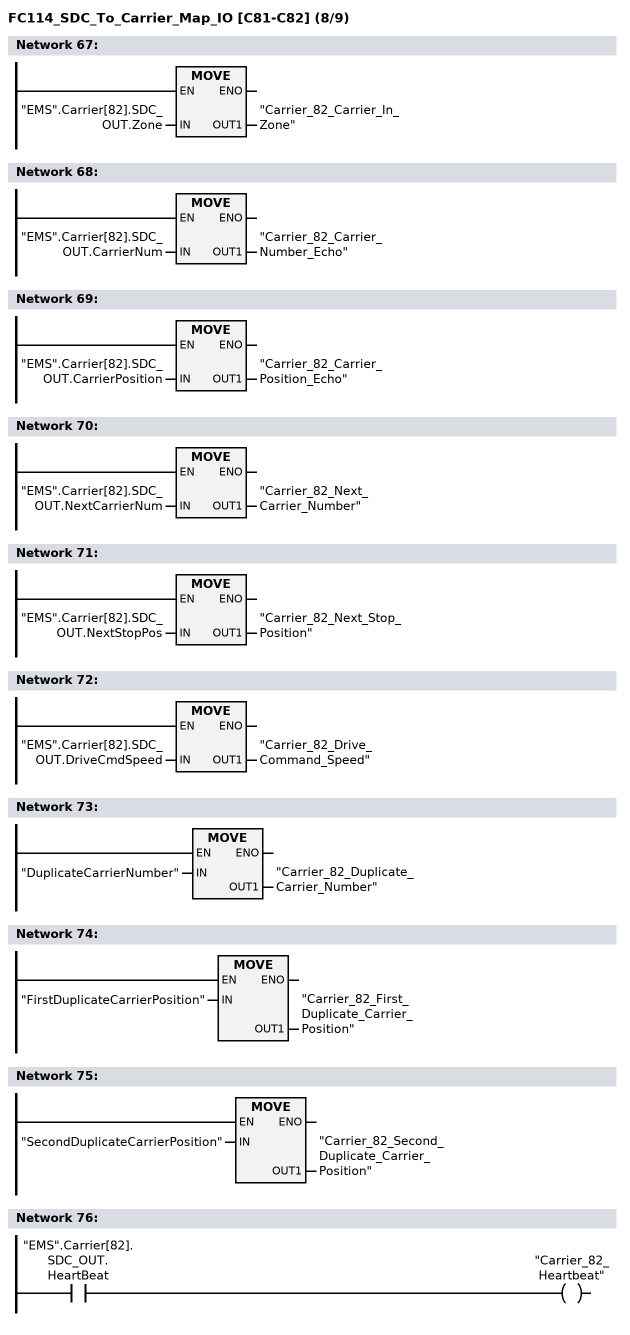
   RUNG wire#powerrail
      Move(in := "EMS".Carrier[82].SDC_OUT.Zone, out1 => "Carrier_82_Carrier_In_Zone")
   END_RUNG
   // the same network as SCL:
   "Carrier_82_Carrier_In_Zone" := "EMS".Carrier[82].SDC_OUT.Zone;
END_REGION

REGION Network 68
   RUNG wire#powerrail
      Move(in := "EMS".Carrier[82].SDC_OUT.CarrierNum, out1 => "Carrier_82_Carrier_Number_Echo")
   END_RUNG
   // the same network as SCL:
   "Carrier_82_Carrier_Number_Echo" := "EMS".Carrier[82].SDC_OUT.CarrierNum;
END_REGION

REGION Network 69
   RUNG wire#powerrail
      Move(in := "EMS".Carrier[82].SDC_OUT.CarrierPosition, out1 => "Carrier_82_Carrier_Position_Echo")
   END_RUNG
   // the same network as SCL:
   "Carrier_82_Carrier_Position_Echo" := "EMS".Carrier[82].SDC_OUT.CarrierPosition;
END_REGION

REGION Network 70
   RUNG wire#powerrail
      Move(in := "EMS".Carrier[82].SDC_OUT.NextCarrierNum, out1 => "Carrier_82_Next_Carrier_Number")
   END_RUNG
   // the same network as SCL:
   "Carrier_82_Next_Carrier_Number" := "EMS".Carrier[82].SDC_OUT.NextCarrierNum;
END_REGION

REGION Network 71
   RUNG wire#powerrail
      Move(in := "EMS".Carrier[82].SDC_OUT.NextStopPos, out1 => "Carrier_82_Next_Stop_Position")
   END_RUNG
   // the same network as SCL:
   "Carrier_82_Next_Stop_Position" := "EMS".Carrier[82].SDC_OUT.NextStopPos;
END_REGION

REGION Network 72
   RUNG wire#powerrail
      Move(in := "EMS".Carrier[82].SDC_OUT.DriveCmdSpeed, out1 => "Carrier_82_Drive_Command_Speed")
   END_RUNG
   // the same network as SCL:
   "Carrier_82_Drive_Command_Speed" := "EMS".Carrier[82].SDC_OUT.DriveCmdSpeed;
END_REGION

REGION Network 73
   RUNG wire#powerrail
      Move(in := "DuplicateCarrierNumber", out1 => "Carrier_82_Duplicate_Carrier_Number")
   END_RUNG
   // the same network as SCL:
   "Carrier_82_Duplicate_Carrier_Number" := "DuplicateCarrierNumber";
END_REGION

REGION Network 74
   RUNG wire#powerrail
      Move(in := "FirstDuplicateCarrierPosition", out1 => "Carrier_82_First_Duplicate_Carrier_Position")
   END_RUNG
   // the same network as SCL:
   "Carrier_82_First_Duplicate_Carrier_Position" := "FirstDuplicateCarrierPosition";
END_REGION

REGION Network 75
   RUNG wire#powerrail
      Move(in := "SecondDuplicateCarrierPosition", out1 => "Carrier_82_Second_Duplicate_Carrier_Position")
   END_RUNG
   // the same network as SCL:
   "Carrier_82_Second_Duplicate_Carrier_Position" := "SecondDuplicateCarrierPosition";
END_REGION

REGION Network 76
   RUNG wire#powerrail
      Contact( "EMS".Carrier[82].SDC_OUT.HeartBeat )
      Coil( "Carrier_82_Heartbeat" )
   END_RUNG
   // the same network as SCL:
   "Carrier_82_Heartbeat" := "EMS".Carrier[82].SDC_OUT.HeartBeat;
END_REGION

REGION Network 77
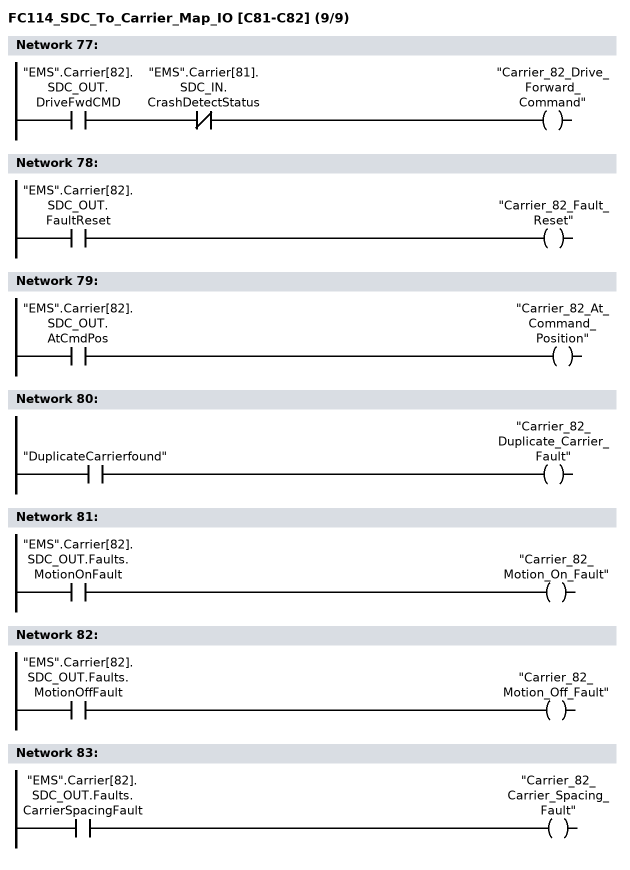
   RUNG wire#powerrail
      Contact( "EMS".Carrier[82].SDC_OUT.DriveFwdCMD )
      I_Contact( "EMS".Carrier[81].SDC_IN.CrashDetectStatus )
      Coil( "Carrier_82_Drive_Forward_Command" )
   END_RUNG
   // the same network as SCL:
   "Carrier_82_Drive_Forward_Command" := "EMS".Carrier[82].SDC_OUT.DriveFwdCMD AND NOT "EMS".Carrier[81].SDC_IN.CrashDetectStatus;
END_REGION

REGION Network 78
   RUNG wire#powerrail
      Contact( "EMS".Carrier[82].SDC_OUT.FaultReset )
      Coil( "Carrier_82_Fault_Reset" )
   END_RUNG
   // the same network as SCL:
   "Carrier_82_Fault_Reset" := "EMS".Carrier[82].SDC_OUT.FaultReset;
END_REGION

REGION Network 79
   RUNG wire#powerrail
      Contact( "EMS".Carrier[82].SDC_OUT.AtCmdPos )
      Coil( "Carrier_82_At_Command_Position" )
   END_RUNG
   // the same network as SCL:
   "Carrier_82_At_Command_Position" := "EMS".Carrier[82].SDC_OUT.AtCmdPos;
END_REGION

REGION Network 80
   RUNG wire#powerrail
      Contact( "DuplicateCarrierfound" )
      Coil( "Carrier_82_Duplicate_Carrier_Fault" )
   END_RUNG
   // the same network as SCL:
   "Carrier_82_Duplicate_Carrier_Fault" := "DuplicateCarrierfound";
END_REGION

REGION Network 81
   RUNG wire#powerrail
      Contact( "EMS".Carrier[82].SDC_OUT.Faults.MotionOnFault )
      Coil( "Carrier_82_Motion_On_Fault" )
   END_RUNG
   // the same network as SCL:
   "Carrier_82_Motion_On_Fault" := "EMS".Carrier[82].SDC_OUT.Faults.MotionOnFault;
END_REGION

REGION Network 82
   RUNG wire#powerrail
      Contact( "EMS".Carrier[82].SDC_OUT.Faults.MotionOffFault )
      Coil( "Carrier_82_Motion_Off_Fault" )
   END_RUNG
   // the same network as SCL:
   "Carrier_82_Motion_Off_Fault" := "EMS".Carrier[82].SDC_OUT.Faults.MotionOffFault;
END_REGION

REGION Network 83
   RUNG wire#powerrail
      Contact( "EMS".Carrier[82].SDC_OUT.Faults.CarrierSpacingFault )
      Coil( "Carrier_82_Carrier_Spacing_Fault" )
   END_RUNG
   // the same network as SCL:
   "Carrier_82_Carrier_Spacing_Fault" := "EMS".Carrier[82].SDC_OUT.Faults.CarrierSpacingFault;
END_REGION
END_FUNCTION

FUNCTION "FC200_FindCarrierZone" : Void   // FC200, SCL
{ S7_Optimized_Access := 'FALSE' }
VERSION : 0.1
   VAR_INPUT
      TotalZones : Int;
      TotalCarriers : Int;
      Reset : Bool;
   END_VAR
   VAR_OUTPUT
      CarrierFindArrayBuffer : "UDT_Carrier";
      DN : Bool;
   END_VAR
   VAR_TEMP
      ZoneCounter : Int;
      ZoneFound : Word;
      CarrierCounter : Int;
      ZouneFound : Int;
   END_VAR
BEGIN
   //[***********************************************************************************NO EDITS*******************************************************************************************************]
   //FC200 - Find Carrier Zone
   //Double loop counter finds which zone carrier is located based on Zone Start Position and End Position and records the result in the system EMS DB for each carrier
   //- EMS.Carrier[x].Zone
   //***************************************************************************************************************************************************************************************************

      #ZoneCounter := 1;
      #CarrierCounter := 1;


       FOR #ZoneCounter := 1 TO #TotalZones DO
           // Statement section FOR
           ;
           WHILE #CarrierCounter <= #TotalCarriers DO
               ;
               IF "EMS".Carrier[#CarrierCounter].Position > "EMS".Zone[#ZoneCounter].StartPos AND
                   "EMS".Carrier[#CarrierCounter].Position < "EMS".Zone[#ZoneCounter].EndPos
                   THEN
                   #CarrierFindArrayBuffer.CARRIER[#CarrierCounter].Zone := #ZoneCounter;
               END_IF;

               #CarrierCounter := #CarrierCounter + 1;
               "cARIERLOOPCOUNT2" := #CarrierCounter;
           END_WHILE;
           #CarrierCounter := 1;
           "ZoneCnt" := #ZoneCounter;
       END_FOR;
END_FUNCTION

FUNCTION "FC201_ZoneCarrierStatus" : Void   // FC201, SCL
{ S7_Optimized_Access := 'FALSE' }
VERSION : 0.1
   VAR_INPUT
      Zone : Int;
      TotalPosition : Int;
      TotalCarriers : Int;
      TotalZones : Int;
      Reset : Bool;
   END_VAR
   VAR_OUTPUT
      ZonePosnArrayBuffer : Array[0..60] of "UDT_ZoneCarrierStatus";
      DN : Bool;
   END_VAR
   VAR_TEMP
      ZoneCounter : Int;
      ZoneFound : Word;
      CarrierCounter : Int;
      SortArrayIndex : Int;
      ArrayIndex : Int;
      Idx1 : Int;
      MaxVal : Int;
      MaxIdx1 : Int;
      Max : Int;
      Idx2 : Int;
      SelectionSort : Int;
   END_VAR
BEGIN
       //[***********************************************************************************NO EDITS*******************************************************************************************************]
       //FC201 - Find Carrier Status
       //Double loop counter finds which zone carrier is located based on Zone Start Position and End Position and records the result in the system EMS DB for each carrier
       //- EMS.Carrier[x].Zone
       //***************************************************************************************************************************************************************************************************

       #CarrierCounter := 1;
       #ArrayIndex := 1;

           WHILE #CarrierCounter <= #TotalCarriers DO
               IF "EMS".Carrier[#CarrierCounter].Zone = #Zone THEN
                   #ZonePosnArrayBuffer[#ArrayIndex].CarrierNumber := "EMS".Carrier[#CarrierCounter].SDC_IN.CarrierNumber;
                   #ZonePosnArrayBuffer[#ArrayIndex].Position := "EMS".Carrier[#CarrierCounter].Position;
                    #ArrayIndex := #ArrayIndex + 1;
                    "IndexArraytemp" := #ArrayIndex;
               ELSE
                   #ZonePosnArrayBuffer[#ArrayIndex].CarrierNumber := 0;
                   #ZonePosnArrayBuffer[#ArrayIndex].Position := 0;
               END_IF;
               #CarrierCounter := #CarrierCounter + 1;
           END_WHILE;
END_FUNCTION

FUNCTION "FC202_ZoneCarrierSort" : Void   // FC202, SCL
{ S7_Optimized_Access := 'FALSE' }
VERSION : 0.1
   VAR_INPUT
      ArrayInUnsort : Array[0..60] of "UDT_ZoneCarrierStatus";
      Max : Int;
   END_VAR
   VAR_OUTPUT
      ZonePositionArrayOut : Array[0..60] of "UDT_ZoneCarrierStatus";
   END_VAR
   VAR_TEMP
      Idx1 : Int;
      MaxVal : DWord;
      MaxIdx1 : Int;
      Idx2 : Int;
      SelectionSort : Int;
      ArrayTemp : Array[0..60] of "UDT_ZoneCarrierStatus";
      MaxCarr : Int;
   END_VAR
BEGIN
   //[***********************************************************************************NO EDITS*******************************************************************************************************]
   //FC202 - Zone Carrier Sort
   //Double loop counter Sorts Carriers in Called Zone to place in correct sequence within  zone. Zones are divided into position based on MaxCarriers allowed in zone as set in the
   //zone setup function block.  Sorted array is used in Traffic cop zone motion control
   //- EMS.Carrier[x].Zone
   //***************************************************************************************************************************************************************************************************
   #ArrayTemp := #ArrayInUnsort;


   FOR #Idx1 := 1 TO #Max BY 1 DO

       #MaxVal := #ArrayTemp[#Idx1].Position;
       IF #ArrayTemp[#Idx1].Position = 0 THEN
           EXIT;
       ELSE
           #MaxIdx1 := #Idx1;
       END_IF;

       FOR #Idx2 := 1 TO #Idx1 + 1 DO
           IF #ArrayTemp[#Idx2].Position > #MaxVal THEN
               #MaxVal := #ArrayTemp[#Idx2].Position;
               #MaxCarr := #ArrayTemp[#Idx2].CarrierNumber;
               #MaxIdx1 := #Idx2;
           END_IF;
       END_FOR;
       IF #MaxIdx1 > #Idx1 THEN
           #ArrayTemp[#MaxIdx1].Position := #ArrayTemp[#Idx1].Position;
           #ArrayTemp[#MaxIdx1].CarrierNumber := #ArrayTemp[#Idx1].CarrierNumber;
           #ArrayTemp[#Idx1].Position := #MaxVal;
           #ArrayTemp[#Idx1].CarrierNumber := #MaxCarr;

       END_IF;

   END_FOR;
   #ZonePositionArrayOut := #ArrayTemp;
END_FUNCTION

FUNCTION "FC203_FindLastZnPos" : Void   // FC203, SCL
{ S7_Optimized_Access := 'FALSE' }
VERSION : 0.1
   VAR_INPUT
      Zone : Int;
      TotalPosition : Int;
   END_VAR
   VAR_OUTPUT
      LastCarrierZnPos : Word;
   END_VAR
   VAR_TEMP
      ZnPosCounter : Int;
      ZoneFound : Word;
      CarrierCounter : Int;
      SortArrayIndex : Int;
      ArrayIndex : Int;
      Idx1 : Int;
      MaxVal : Int;
      MaxIdx1 : Int;
      Max : Int;
      Idx2 : Int;
      SelectionSort : Int;
   END_VAR
BEGIN
       #ZnPosCounter := #TotalPosition;
       WHILE #ZnPosCounter >= 1 DO

           IF "EMS".Zone[#Zone].CarrierZnStatus[#ZnPosCounter].CarrierNumber <> 0 THEN
               ;
               #LastCarrierZnPos := #ZnPosCounter;
               RETURN;
           END_IF;
           #ZnPosCounter := #ZnPosCounter - 1;
       END_WHILE;
END_FUNCTION

FUNCTION "FC204_FindCarrierZNPos" : Void   // FC204, SCL
{ S7_Optimized_Access := 'FALSE' }
VERSION : 0.1
   VAR_INPUT
      Carrier : Word;
      Zone : Int;
      TotalPosition : Int;
   END_VAR
   VAR_OUTPUT
      CarrierZnPos : Word;
   END_VAR
   VAR_TEMP
      ZnPosCounter : Int;
      ZoneFound : Word;
      CarrierCounter : Int;
      SortArrayIndex : Int;
      ArrayIndex : Int;
      Idx1 : Int;
      MaxVal : Int;
      MaxIdx1 : Int;
      Max : Int;
      Idx2 : Int;
      SelectionSort : Int;
   END_VAR
BEGIN
   //[***********************************************************************************NO EDITS*******************************************************************************************************]
   //FC204 - Find Carrier Zone Position
   //Single loop Counter finds which #Zone Position. Zone Position is determined BY Value OF Max Carriers defined in  #Carrier is located based on #Zone Start Position AND End Position AND
   //records the result in the system "EMS" DB FOR each Zone and the results stored in the EMS.Zone[Zone].CarrierZnStatus[1 thru Max Carriers in Zone].Carrier Number
   //***************************************************************************************************************************************************************************************************   

       #ZnPosCounter := 1;
       FOR #ZnPosCounter := 1 TO #TotalPosition DO
           ;
           IF "EMS".Zone[#Zone].CarrierZnStatus[#ZnPosCounter].CarrierNumber = #Carrier THEN;
               ;
               #CarrierZnPos := #ZnPosCounter;
           END_IF;
       END_FOR;
END_FUNCTION

FUNCTION "FC205_FindDuplicateCarrier" : Void   // FC205, SCL
{ S7_Optimized_Access := 'TRUE' }
VERSION : 0.1
   VAR_INPUT
      Carrier : Array[0..99] of "UDT_CarrierStructure";
      TotalCarriers : Int;
   END_VAR
   VAR_OUTPUT
      DuplicateFound : Bool;
      DuplicateCarrierNumber : Word;
      FirstDuplicatePosition : Word;
      SecondDuplicate : Word;
   END_VAR
   VAR_TEMP
      CarrierFindCnt : Int;
      temp1 : Int;
      CarrierCounter : Int;
      CarrierFindArray : Array[0..99] of "UDT_CarrierStructure";
   END_VAR
BEGIN
   //Sorts Carriers in Called Zone TO place in correct sequence within  Zone. Zones are divided into position based on MaxCarriers allowed in Zone as set in the Zone setup function block.


   #DuplicateFound := FALSE;
   #CarrierCounter := 1;
   #CarrierFindCnt := 1;
   #CarrierFindArray := #Carrier;
   FOR #CarrierFindCnt := 1 TO #TotalCarriers DO
       ;
       WHILE #CarrierCounter <= #TotalCarriers DO
           ;
           IF #Carrier[#CarrierCounter].SDC_IN.CarrierNumber = #CarrierFindArray[#CarrierFindCnt].SDC_IN.CarrierNumber AND #CarrierCounter <> #CarrierFindCnt AND #Carrier[#CarrierCounter].SDC_IN.CarrierNumber <> 0 THEN
               #DuplicateFound := TRUE;
               #FirstDuplicatePosition:= #Carrier[#CarrierCounter].SDC_IN.CarrierPosition;
               #SecondDuplicate := #Carrier[#CarrierFindCnt].SDC_IN.CarrierPosition;
               #DuplicateCarrierNumber := #CarrierFindArray[#CarrierFindCnt].SDC_IN.CarrierNumber;
               RETURN;
           END_IF;
           #CarrierCounter := #CarrierCounter + 1;
       END_WHILE;

       #CarrierCounter := 1;
   END_FOR;
END_FUNCTION

FUNCTION "FC206_HMIZonePosTracking" : Void   // FC206, SCL
{ S7_Optimized_Access := 'FALSE' }
VERSION : 0.1
   VAR_INPUT
      Zone : Int;
      TotalZones : Int;
      TotalCarriers : Int;
      MaxCarrierPosns : Int;
   END_VAR
   VAR_OUTPUT
      HMIZonePositionDisplay : Array[1..20] of "UDT_HMIZonePositionStructure";
   END_VAR
   VAR_TEMP
      PositionCounter : Int;
      ZoneFound : Word;
      CarrierCounter : Int;
      ZouneFound : Int;
   END_VAR
BEGIN

       FOR #PositionCounter := 1 TO #MaxCarrierPosns BY 1 DO
           FOR #CarrierCounter := 1 TO #TotalCarriers BY 1 DO
               ;
               IF "EMS".Carrier[#CarrierCounter].Position >= "EMS".Zone[#Zone].HMIZonePositions[#PositionCounter].ZonePosition AND
                   "EMS".Carrier[#CarrierCounter].Position < "EMS".Zone[#Zone].HMIZonePositions[#PositionCounter + 1].ZonePosition
               THEN
                   #HMIZonePositionDisplay[#PositionCounter].CarrierNumber := #CarrierCounter;
                   #HMIZonePositionDisplay[#PositionCounter].CarrierPosition := "EMS".Carrier[#CarrierCounter].Position;
                   #HMIZonePositionDisplay[#PositionCounter].Faulted := "EMS".Carrier[#CarrierCounter].Faulted;
                   EXIT;
               ELSE
                   ;
                   #HMIZonePositionDisplay[#PositionCounter].CarrierNumber := 0;
                   #HMIZonePositionDisplay[#PositionCounter].CarrierPosition := 0;
                   #HMIZonePositionDisplay[#PositionCounter].Faulted := 0;
               END_IF;
               "FC206CarrierLoop" := #CarrierCounter;
           END_FOR;
       "FC206PositionLoop" := #PositionCounter;
   END_FOR;
END_FUNCTION

FUNCTION "FC301_StopZone1_TrafficCop" : Void   // FC301, LAD
{ S7_Optimized_Access := 'TRUE' }
VERSION : 0.1
   VAR_INPUT
      Zone : Int;
   END_VAR
   VAR_TEMP
      TrafficCopCarrier : Int;
      CarrierMotionZn : Array[0..40] of "UDT_ZoneCarrierStatus";
      InTransitMemory : Bool;
   END_VAR
BEGIN

REGION Network 1
   // **********************************************************************************************************************
   // 
   // Zone Function Block.  Static setup of all Zone Parameters.  Traffic Cop Setup Logic - Handles all motion and carrier movement logic based on interdependence of Each Carrier in Zone # Passed from Main program Call in OB1 
   // 
   // **********************************************************************************************************************
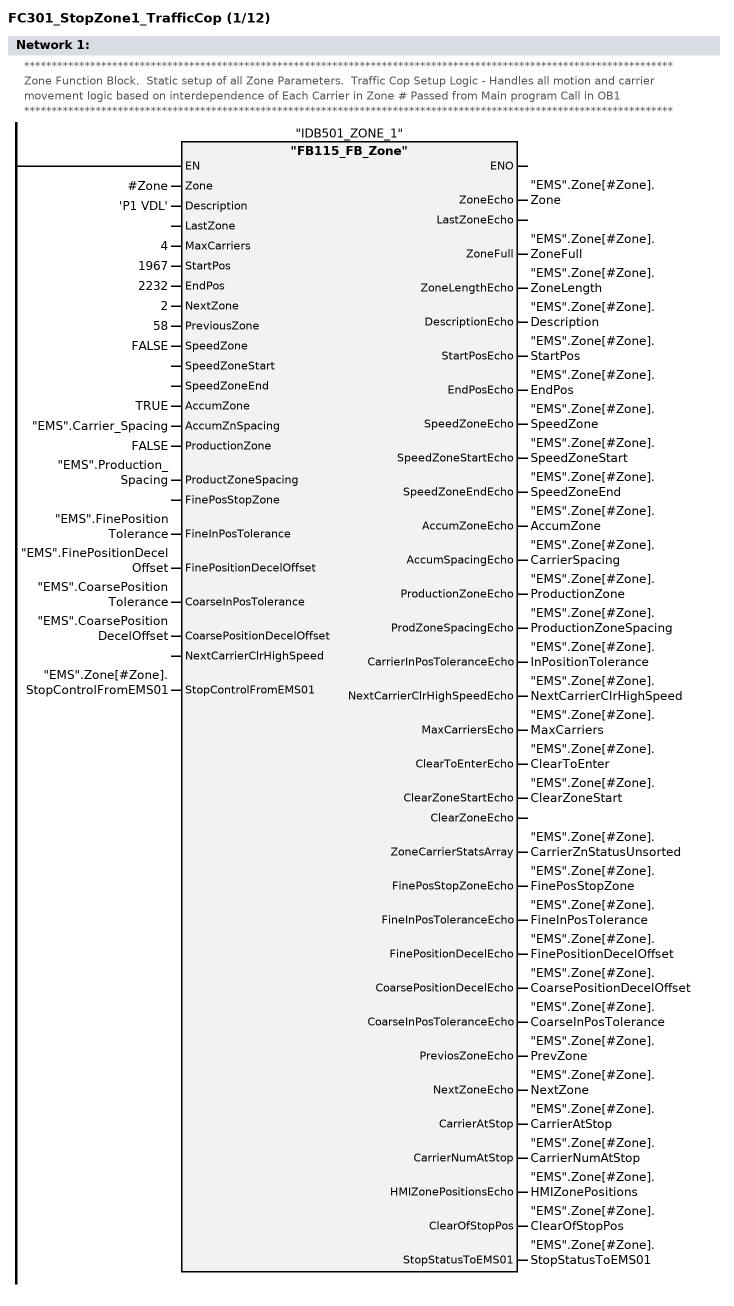
   RUNG wire#powerrail
      "IDB501_ZONE_1"(Zone := #Zone, Description := 'P1 VDL', LastZone :=, MaxCarriers := 4, StartPos := 1967, EndPos := 2232, NextZone := 2, PreviousZone := 58, SpeedZone := FALSE, SpeedZoneStart :=, SpeedZoneEnd :=, AccumZone := TRUE, AccumZnSpacing := "EMS".Carrier_Spacing, ProductionZone := FALSE, ProductZoneSpacing := "EMS".Production_Spacing, FinePosStopZone :=, FineInPosTolerance := "EMS".FinePositionTolerance, FinePositionDecelOffset := "EMS".FinePositionDecelOffset, CoarseInPosTolerance := "EMS".CoarsePositionTolerance, CoarsePositionDecelOffset := "EMS".CoarsePositionDecelOffset, NextCarrierClrHighSpeed :=, StopControlFromEMS01 := "EMS".Zone[#Zone].StopControlFromEMS01, ZoneEcho => "EMS".Zone[#Zone].Zone, LastZoneEcho =>, ZoneFull => "EMS".Zone[#Zone].ZoneFull, ZoneLengthEcho => "EMS".Zone[#Zone].ZoneLength, DescriptionEcho => "EMS".Zone[#Zone].Description, StartPosEcho => "EMS".Zone[#Zone].StartPos, EndPosEcho => "EMS".Zone[#Zone].EndPos, SpeedZoneEcho => "EMS".Zone[#Zone].SpeedZone, SpeedZoneStartEcho => "EMS".Zone[#Zone].SpeedZoneStart, SpeedZoneEndEcho => "EMS".Zone[#Zone].SpeedZoneEnd, AccumZoneEcho => "EMS".Zone[#Zone].AccumZone, AccumSpacingEcho => "EMS".Zone[#Zone].CarrierSpacing, ProductionZoneEcho => "EMS".Zone[#Zone].ProductionZone, ProdZoneSpacingEcho => "EMS".Zone[#Zone].ProductionZoneSpacing, CarrierInPosToleranceEcho => "EMS".Zone[#Zone].InPositionTolerance, NextCarrierClrHighSpeedEcho => "EMS".Zone[#Zone].NextCarrierClrHighSpeed, MaxCarriersEcho => "EMS".Zone[#Zone].MaxCarriers, ClearToEnterEcho => "EMS".Zone[#Zone].ClearToEnter, ClearZoneStartEcho => "EMS".Zone[#Zone].ClearZoneStart, ClearZoneEcho =>, ZoneCarrierStatsArray => "EMS".Zone[#Zone].CarrierZnStatusUnsorted, FinePosStopZoneEcho => "EMS".Zone[#Zone].FinePosStopZone, FineInPosToleranceEcho => "EMS".Zone[#Zone].FineInPosTolerance, FinePositionDecelEcho => "EMS".Zone[#Zone].FinePositionDecelOffset, CoarsePositionDecelEcho => "EMS".Zone[#Zone].CoarsePositionDecelOffset, CoarseInPosToleranceEcho => "EMS".Zone[#Zone].CoarseInPosTolerance, PreviosZoneEcho => "EMS".Zone[#Zone].PrevZone, NextZoneEcho => "EMS".Zone[#Zone].NextZone, CarrierAtStop => "EMS".Zone[#Zone].CarrierAtStop, CarrierNumAtStop => "EMS".Zone[#Zone].CarrierNumAtStop, HMIZonePositionsEcho => "EMS".Zone[#Zone].HMIZonePositions, ClearOfStopPos => "EMS".Zone[#Zone].ClearOfStopPos, StopStatusToEMS01 => "EMS".Zone[#Zone].StopStatusToEMS01)
   END_RUNG
   // the same network as SCL:
   "IDB501_ZONE_1"(Zone := #Zone,   // "FB115_FB_Zone"
                   Description := 'P1 VDL',
                   MaxCarriers := 4,
                   StartPos := 1967,
                   EndPos := 2232,
                   NextZone := 2,
                   PreviousZone := 58,
                   SpeedZone := FALSE,
                   AccumZone := TRUE,
                   AccumZnSpacing := "EMS".Carrier_Spacing,
                   ProductionZone := FALSE,
                   ProductZoneSpacing := "EMS".Production_Spacing,
                   FineInPosTolerance := "EMS".FinePositionTolerance,
                   FinePositionDecelOffset := "EMS".FinePositionDecelOffset,
                   CoarseInPosTolerance := "EMS".CoarsePositionTolerance,
                   CoarsePositionDecelOffset := "EMS".CoarsePositionDecelOffset,
                   StopControlFromEMS01 := "EMS".Zone[#Zone].StopControlFromEMS01,
                   ZoneEcho => "EMS".Zone[#Zone].Zone,
                   ZoneFull => "EMS".Zone[#Zone].ZoneFull,
                   ZoneLengthEcho => "EMS".Zone[#Zone].ZoneLength,
                   DescriptionEcho => "EMS".Zone[#Zone].Description,
                   StartPosEcho => "EMS".Zone[#Zone].StartPos,
                   EndPosEcho => "EMS".Zone[#Zone].EndPos,
                   SpeedZoneEcho => "EMS".Zone[#Zone].SpeedZone,
                   SpeedZoneStartEcho => "EMS".Zone[#Zone].SpeedZoneStart,
                   SpeedZoneEndEcho => "EMS".Zone[#Zone].SpeedZoneEnd,
                   AccumZoneEcho => "EMS".Zone[#Zone].AccumZone,
                   AccumSpacingEcho => "EMS".Zone[#Zone].CarrierSpacing,
                   ProductionZoneEcho => "EMS".Zone[#Zone].ProductionZone,
                   ProdZoneSpacingEcho => "EMS".Zone[#Zone].ProductionZoneSpacing,
                   CarrierInPosToleranceEcho => "EMS".Zone[#Zone].InPositionTolerance,
                   NextCarrierClrHighSpeedEcho => "EMS".Zone[#Zone].NextCarrierClrHighSpeed,
                   MaxCarriersEcho => "EMS".Zone[#Zone].MaxCarriers,
                   ClearToEnterEcho => "EMS".Zone[#Zone].ClearToEnter,
                   ClearZoneStartEcho => "EMS".Zone[#Zone].ClearZoneStart,
                   ZoneCarrierStatsArray => "EMS".Zone[#Zone].CarrierZnStatusUnsorted,
                   FinePosStopZoneEcho => "EMS".Zone[#Zone].FinePosStopZone,
                   FineInPosToleranceEcho => "EMS".Zone[#Zone].FineInPosTolerance,
                   FinePositionDecelEcho => "EMS".Zone[#Zone].FinePositionDecelOffset,
                   CoarsePositionDecelEcho => "EMS".Zone[#Zone].CoarsePositionDecelOffset,
                   CoarseInPosToleranceEcho => "EMS".Zone[#Zone].CoarseInPosTolerance,
                   PreviosZoneEcho => "EMS".Zone[#Zone].PrevZone,
                   NextZoneEcho => "EMS".Zone[#Zone].NextZone,
                   CarrierAtStop => "EMS".Zone[#Zone].CarrierAtStop,
                   CarrierNumAtStop => "EMS".Zone[#Zone].CarrierNumAtStop,
                   HMIZonePositionsEcho => "EMS".Zone[#Zone].HMIZonePositions,
                   ClearOfStopPos => "EMS".Zone[#Zone].ClearOfStopPos,
                   StopStatusToEMS01 => "EMS".Zone[#Zone].StopStatusToEMS01);
END_REGION

REGION Network 2
   // *********************************************************************************************************************
   // Carrier Sort Function FC202 - Sorts Carriers in Called Zone to place in correct sequence within  zone. Zones are divided into position based on MaxCarriers allowed in zone as set in the zone setup function block. 
   // 
   // **********************************************************************************************************************
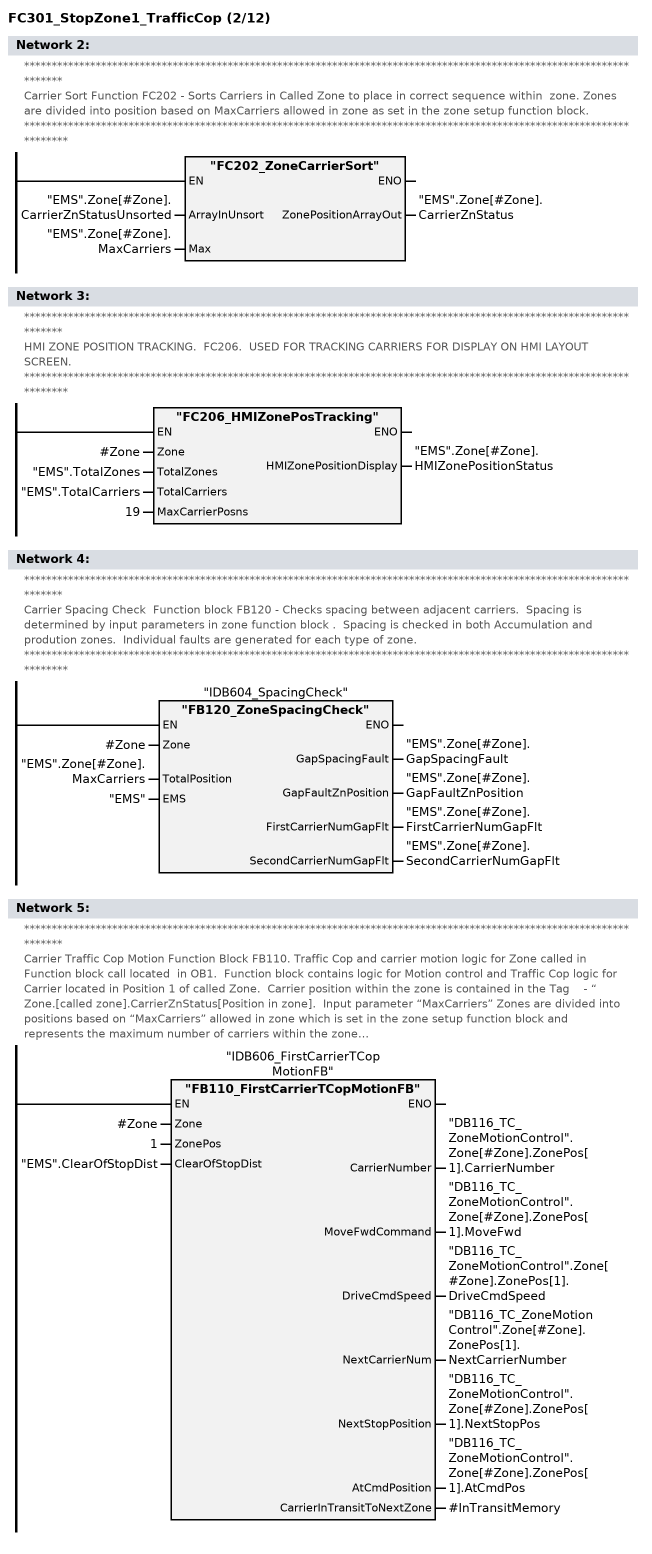
   RUNG wire#powerrail
      "FC202_ZoneCarrierSort"(ArrayInUnsort := "EMS".Zone[#Zone].CarrierZnStatusUnsorted, Max := "EMS".Zone[#Zone].MaxCarriers, ZonePositionArrayOut => "EMS".Zone[#Zone].CarrierZnStatus)
   END_RUNG
   // the same network as SCL:
   "FC202_ZoneCarrierSort"(ArrayInUnsort := "EMS".Zone[#Zone].CarrierZnStatusUnsorted,
                           Max := "EMS".Zone[#Zone].MaxCarriers,
                           ZonePositionArrayOut => "EMS".Zone[#Zone].CarrierZnStatus);
END_REGION

REGION Network 3
   // *********************************************************************************************************************
   // HMI ZONE POSITION TRACKING.  FC206.  USED FOR TRACKING CARRIERS FOR DISPLAY ON HMI LAYOUT SCREEN. 
   // **********************************************************************************************************************
   RUNG wire#powerrail
      "FC206_HMIZonePosTracking"(Zone := #Zone, TotalZones := "EMS".TotalZones, TotalCarriers := "EMS".TotalCarriers, MaxCarrierPosns := 19, HMIZonePositionDisplay => "EMS".Zone[#Zone].HMIZonePositionStatus)
   END_RUNG
   // the same network as SCL:
   "FC206_HMIZonePosTracking"(Zone := #Zone,
                           TotalZones := "EMS".TotalZones,
                           TotalCarriers := "EMS".TotalCarriers,
                           MaxCarrierPosns := 19,
                           HMIZonePositionDisplay => "EMS".Zone[#Zone].HMIZonePositionStatus);
END_REGION

REGION Network 4
   // *********************************************************************************************************************
   // 
   // Carrier Spacing Check  Function block FB120 - Checks spacing between adjacent carriers.  Spacing is determined by input parameters in zone function block .  Spacing is checked in both Accumulation and prodution zones.  Individual faults are generated for each type of zone.
   // 
   // **********************************************************************************************************************
   RUNG wire#powerrail
      "IDB604_SpacingCheck"(Zone := #Zone, TotalPosition := "EMS".Zone[#Zone].MaxCarriers, EMS := "EMS", GapSpacingFault => "EMS".Zone[#Zone].GapSpacingFault, GapFaultZnPosition => "EMS".Zone[#Zone].GapFaultZnPosition, FirstCarrierNumGapFlt => "EMS".Zone[#Zone].FirstCarrierNumGapFlt, SecondCarrierNumGapFlt => "EMS".Zone[#Zone].SecondCarrierNumGapFlt)
   END_RUNG
   // the same network as SCL:
   "IDB604_SpacingCheck"(Zone := #Zone,   // "FB120_ZoneSpacingCheck"
                         TotalPosition := "EMS".Zone[#Zone].MaxCarriers,
                         EMS := "EMS",
                         GapSpacingFault => "EMS".Zone[#Zone].GapSpacingFault,
                         GapFaultZnPosition => "EMS".Zone[#Zone].GapFaultZnPosition,
                         FirstCarrierNumGapFlt => "EMS".Zone[#Zone].FirstCarrierNumGapFlt,
                         SecondCarrierNumGapFlt => "EMS".Zone[#Zone].SecondCarrierNumGapFlt);
END_REGION

REGION Network 5
   // *********************************************************************************************************************
   // 
   // Carrier Traffic Cop Motion Function Block FB110. Traffic Cop and carrier motion logic for Zone called in Function block call located  in OB1.  Function block contains logic for Motion control and Traffic Cop logic for Carrier located in Position 1 of called Zone.  Carrier position within the zone is contained in the Tag    - “ Zone.[called zone].CarrierZnStatus[Position in zone].  Input parameter “MaxCarriers” Zones are divided into positions based on “MaxCarriers” allowed in zone which is set in the zone setup function block and represents the maximum number of carriers within the zone. 
   // 
   // **********************************************************************************************************************
   RUNG wire#powerrail
      "IDB606_FirstCarrierTCopMotionFB"(Zone := #Zone, ZonePos := 1, ClearOfStopDist := "EMS".ClearOfStopDist, CarrierNumber => "DB116_TC_ZoneMotionControl".Zone[#Zone].ZonePos[1].CarrierNumber, MoveFwdCommand => "DB116_TC_ZoneMotionControl".Zone[#Zone].ZonePos[1].MoveFwd, DriveCmdSpeed => "DB116_TC_ZoneMotionControl".Zone[#Zone].ZonePos[1].DriveCmdSpeed, NextCarrierNum => "DB116_TC_ZoneMotionControl".Zone[#Zone].ZonePos[1].NextCarrierNumber, NextStopPosition => "DB116_TC_ZoneMotionControl".Zone[#Zone].ZonePos[1].NextStopPos, AtCmdPosition => "DB116_TC_ZoneMotionControl".Zone[#Zone].ZonePos[1].AtCmdPos, CarrierInTransitToNextZone => #InTransitMemory)
   END_RUNG
   // the same network as SCL:
   "IDB606_FirstCarrierTCopMotionFB"(Zone := #Zone,   // "FB110_FirstCarrierTCopMotionFB"
                           ZonePos := 1,
                           ClearOfStopDist := "EMS".ClearOfStopDist,
                           CarrierNumber => "DB116_TC_ZoneMotionControl".Zone[#Zone].ZonePos[1].CarrierNumber,
                           MoveFwdCommand => "DB116_TC_ZoneMotionControl".Zone[#Zone].ZonePos[1].MoveFwd,
                           DriveCmdSpeed => "DB116_TC_ZoneMotionControl".Zone[#Zone].ZonePos[1].DriveCmdSpeed,
                           NextCarrierNum => "DB116_TC_ZoneMotionControl".Zone[#Zone].ZonePos[1].NextCarrierNumber,
                           NextStopPosition => "DB116_TC_ZoneMotionControl".Zone[#Zone].ZonePos[1].NextStopPos,
                           AtCmdPosition => "DB116_TC_ZoneMotionControl".Zone[#Zone].ZonePos[1].AtCmdPos,
                           CarrierInTransitToNextZone => #InTransitMemory);
END_REGION

REGION Network 6
   // *********************************************************************************************************************
   // 
   // Carrier Traffic Cop Motion Function Block FB111. Traffic Cop and carrier motion logic for Zone called in Function block call located  in OB1.  Function block contains logic for Motion control and Traffic Cop logic for Carrier located in Position 2 to the last carrier of called Zone.  Carrier position within the zone is contained in the Tag    - “ Zone.[called zone].CarrierZnStatus[Position in zone].  Input parameter “MaxCarriers” Zones are divided into positions based on “MaxCarriers” allowed in zone which is set in the zone setup function block and represents the maximum number of carriers within the zone. 
   // 
   // **********************************************************************************************************************
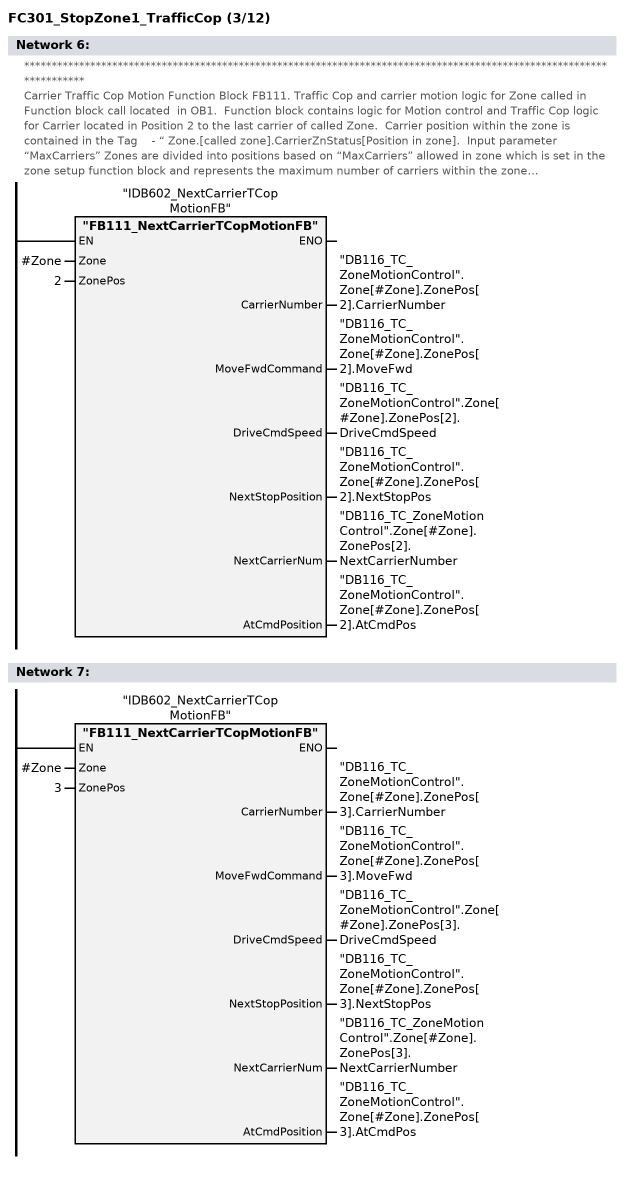
   RUNG wire#powerrail
      "IDB602_NextCarrierTCopMotionFB"(Zone := #Zone, ZonePos := 2, CarrierNumber => "DB116_TC_ZoneMotionControl".Zone[#Zone].ZonePos[2].CarrierNumber, MoveFwdCommand => "DB116_TC_ZoneMotionControl".Zone[#Zone].ZonePos[2].MoveFwd, DriveCmdSpeed => "DB116_TC_ZoneMotionControl".Zone[#Zone].ZonePos[2].DriveCmdSpeed, NextStopPosition => "DB116_TC_ZoneMotionControl".Zone[#Zone].ZonePos[2].NextStopPos, NextCarrierNum => "DB116_TC_ZoneMotionControl".Zone[#Zone].ZonePos[2].NextCarrierNumber, AtCmdPosition => "DB116_TC_ZoneMotionControl".Zone[#Zone].ZonePos[2].AtCmdPos)
   END_RUNG
   // the same network as SCL:
   "IDB602_NextCarrierTCopMotionFB"(Zone := #Zone,   // "FB111_NextCarrierTCopMotionFB"
                           ZonePos := 2,
                           CarrierNumber => "DB116_TC_ZoneMotionControl".Zone[#Zone].ZonePos[2].CarrierNumber,
                           MoveFwdCommand => "DB116_TC_ZoneMotionControl".Zone[#Zone].ZonePos[2].MoveFwd,
                           DriveCmdSpeed => "DB116_TC_ZoneMotionControl".Zone[#Zone].ZonePos[2].DriveCmdSpeed,
                           NextStopPosition => "DB116_TC_ZoneMotionControl".Zone[#Zone].ZonePos[2].NextStopPos,
                           NextCarrierNum => "DB116_TC_ZoneMotionControl".Zone[#Zone].ZonePos[2].NextCarrierNumber,
                           AtCmdPosition => "DB116_TC_ZoneMotionControl".Zone[#Zone].ZonePos[2].AtCmdPos);
END_REGION

REGION Network 7
   RUNG wire#powerrail
      "IDB602_NextCarrierTCopMotionFB"(Zone := #Zone, ZonePos := 3, CarrierNumber => "DB116_TC_ZoneMotionControl".Zone[#Zone].ZonePos[3].CarrierNumber, MoveFwdCommand => "DB116_TC_ZoneMotionControl".Zone[#Zone].ZonePos[3].MoveFwd, DriveCmdSpeed => "DB116_TC_ZoneMotionControl".Zone[#Zone].ZonePos[3].DriveCmdSpeed, NextStopPosition => "DB116_TC_ZoneMotionControl".Zone[#Zone].ZonePos[3].NextStopPos, NextCarrierNum => "DB116_TC_ZoneMotionControl".Zone[#Zone].ZonePos[3].NextCarrierNumber, AtCmdPosition => "DB116_TC_ZoneMotionControl".Zone[#Zone].ZonePos[3].AtCmdPos)
   END_RUNG
   // the same network as SCL:
   "IDB602_NextCarrierTCopMotionFB"(Zone := #Zone,   // "FB111_NextCarrierTCopMotionFB"
                           ZonePos := 3,
                           CarrierNumber => "DB116_TC_ZoneMotionControl".Zone[#Zone].ZonePos[3].CarrierNumber,
                           MoveFwdCommand => "DB116_TC_ZoneMotionControl".Zone[#Zone].ZonePos[3].MoveFwd,
                           DriveCmdSpeed => "DB116_TC_ZoneMotionControl".Zone[#Zone].ZonePos[3].DriveCmdSpeed,
                           NextStopPosition => "DB116_TC_ZoneMotionControl".Zone[#Zone].ZonePos[3].NextStopPos,
                           NextCarrierNum => "DB116_TC_ZoneMotionControl".Zone[#Zone].ZonePos[3].NextCarrierNumber,
                           AtCmdPosition => "DB116_TC_ZoneMotionControl".Zone[#Zone].ZonePos[3].AtCmdPos);
END_REGION

REGION Network 8
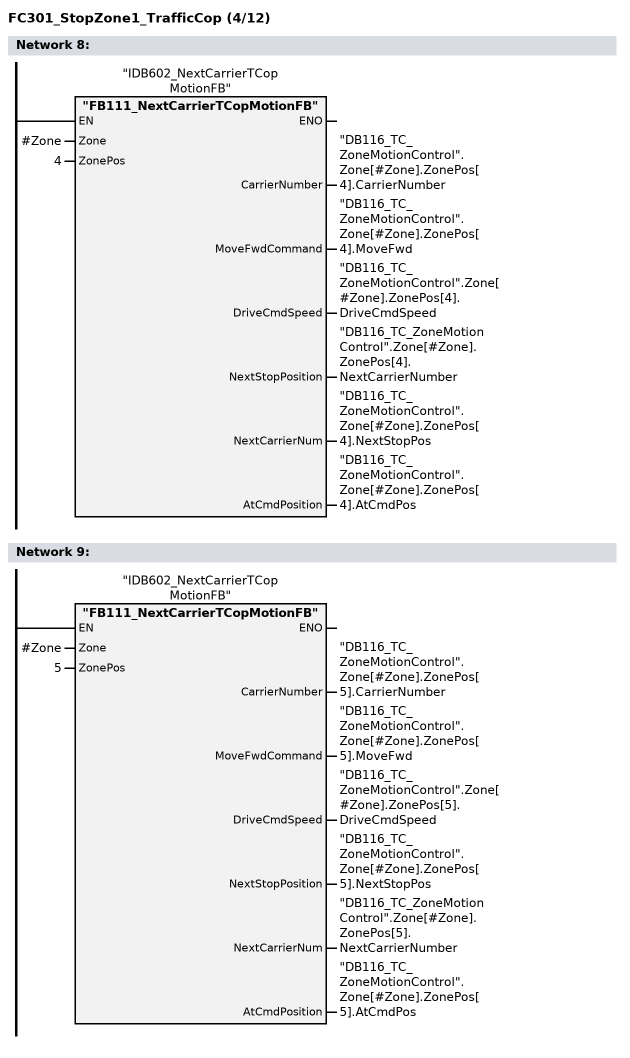
   RUNG wire#powerrail
      "IDB602_NextCarrierTCopMotionFB"(Zone := #Zone, ZonePos := 4, CarrierNumber => "DB116_TC_ZoneMotionControl".Zone[#Zone].ZonePos[4].CarrierNumber, MoveFwdCommand => "DB116_TC_ZoneMotionControl".Zone[#Zone].ZonePos[4].MoveFwd, DriveCmdSpeed => "DB116_TC_ZoneMotionControl".Zone[#Zone].ZonePos[4].DriveCmdSpeed, NextStopPosition => "DB116_TC_ZoneMotionControl".Zone[#Zone].ZonePos[4].NextCarrierNumber, NextCarrierNum => "DB116_TC_ZoneMotionControl".Zone[#Zone].ZonePos[4].NextStopPos, AtCmdPosition => "DB116_TC_ZoneMotionControl".Zone[#Zone].ZonePos[4].AtCmdPos)
   END_RUNG
   // the same network as SCL:
   "IDB602_NextCarrierTCopMotionFB"(Zone := #Zone,   // "FB111_NextCarrierTCopMotionFB"
                           ZonePos := 4,
                           CarrierNumber => "DB116_TC_ZoneMotionControl".Zone[#Zone].ZonePos[4].CarrierNumber,
                           MoveFwdCommand => "DB116_TC_ZoneMotionControl".Zone[#Zone].ZonePos[4].MoveFwd,
                           DriveCmdSpeed => "DB116_TC_ZoneMotionControl".Zone[#Zone].ZonePos[4].DriveCmdSpeed,
                           NextStopPosition => "DB116_TC_ZoneMotionControl".Zone[#Zone].ZonePos[4].NextCarrierNumber,
                           NextCarrierNum => "DB116_TC_ZoneMotionControl".Zone[#Zone].ZonePos[4].NextStopPos,
                           AtCmdPosition => "DB116_TC_ZoneMotionControl".Zone[#Zone].ZonePos[4].AtCmdPos);
END_REGION

REGION Network 9
   RUNG wire#powerrail
      "IDB602_NextCarrierTCopMotionFB"(Zone := #Zone, ZonePos := 5, CarrierNumber => "DB116_TC_ZoneMotionControl".Zone[#Zone].ZonePos[5].CarrierNumber, MoveFwdCommand => "DB116_TC_ZoneMotionControl".Zone[#Zone].ZonePos[5].MoveFwd, DriveCmdSpeed => "DB116_TC_ZoneMotionControl".Zone[#Zone].ZonePos[5].DriveCmdSpeed, NextStopPosition => "DB116_TC_ZoneMotionControl".Zone[#Zone].ZonePos[5].NextStopPos, NextCarrierNum => "DB116_TC_ZoneMotionControl".Zone[#Zone].ZonePos[5].NextCarrierNumber, AtCmdPosition => "DB116_TC_ZoneMotionControl".Zone[#Zone].ZonePos[5].AtCmdPos)
   END_RUNG
   // the same network as SCL:
   "IDB602_NextCarrierTCopMotionFB"(Zone := #Zone,   // "FB111_NextCarrierTCopMotionFB"
                           ZonePos := 5,
                           CarrierNumber => "DB116_TC_ZoneMotionControl".Zone[#Zone].ZonePos[5].CarrierNumber,
                           MoveFwdCommand => "DB116_TC_ZoneMotionControl".Zone[#Zone].ZonePos[5].MoveFwd,
                           DriveCmdSpeed => "DB116_TC_ZoneMotionControl".Zone[#Zone].ZonePos[5].DriveCmdSpeed,
                           NextStopPosition => "DB116_TC_ZoneMotionControl".Zone[#Zone].ZonePos[5].NextStopPos,
                           NextCarrierNum => "DB116_TC_ZoneMotionControl".Zone[#Zone].ZonePos[5].NextCarrierNumber,
                           AtCmdPosition => "DB116_TC_ZoneMotionControl".Zone[#Zone].ZonePos[5].AtCmdPos);
END_REGION

REGION Network 10
